REGION Network 8: WLAN5 Comm Fault
   RUNG wire#powerrail
      Contact( "reset" )
      { S7_Templates := "SrcType := USInt" } EQ_Contact(in1 := "UserDiag_HmiData".actIOSystemData.actIODeviceState[105], in2 := 3)
      wire#w1
      Coil( "DB302_HMI_Faults".SDC_Faults_0.%X5 )
   END_RUNG
   RUNG wire#powerrail
      Contact( "DB302_HMI_Faults".SDC_Faults_0.%X5 )
      I_Contact( "EMS_Fault_Reset" )
   END_RUNG wire#w1
   RUNG wire#w1
      Move(in := 6, out1 => "DB101_DB_SDC_FAULTS".SDC_Fault)
   END_RUNG
   // the same network as SCL:
   "DB302_HMI_Faults".SDC_Faults_0.%X5 := ("reset" AND ("UserDiag_HmiData".actIOSystemData.actIODeviceState[105] = 3)) OR ("DB302_HMI_Faults".SDC_Faults_0.%X5 AND NOT "EMS_Fault_Reset");
   IF "DB302_HMI_Faults".SDC_Faults_0.%X5 THEN "DB101_DB_SDC_FAULTS".SDC_Fault := 6; END_IF;
END_REGION

REGION Network 9: WLAN6 Comm Fault
   RUNG wire#powerrail
      Contact( "reset" )
      { S7_Templates := "SrcType := USInt" } EQ_Contact(in1 := "UserDiag_HmiData".actIOSystemData.actIODeviceState[106], in2 := 3)
      wire#w1
      Coil( "DB302_HMI_Faults".SDC_Faults_0.%X6 )
   END_RUNG
   RUNG wire#powerrail
      Contact( "DB302_HMI_Faults".SDC_Faults_0.%X6 )
      I_Contact( "EMS_Fault_Reset" )
   END_RUNG wire#w1
   RUNG wire#w1
      Move(in := 7, out1 => "DB101_DB_SDC_FAULTS".SDC_Fault)
   END_RUNG
   // the same network as SCL:
   "DB302_HMI_Faults".SDC_Faults_0.%X6 := ("reset" AND ("UserDiag_HmiData".actIOSystemData.actIODeviceState[106] = 3)) OR ("DB302_HMI_Faults".SDC_Faults_0.%X6 AND NOT "EMS_Fault_Reset");
   IF "DB302_HMI_Faults".SDC_Faults_0.%X6 THEN "DB101_DB_SDC_FAULTS".SDC_Fault := 7; END_IF;
END_REGION

REGION Network 10: WLAN7 Comm Fault
   RUNG wire#powerrail
      Contact( "reset" )
      { S7_Templates := "SrcType := USInt" } EQ_Contact(in1 := "UserDiag_HmiData".actIOSystemData.actIODeviceState[107], in2 := 3)
      wire#w1
      Coil( "DB302_HMI_Faults".SDC_Faults_0.%X7 )
   END_RUNG
   RUNG wire#powerrail
      Contact( "DB302_HMI_Faults".SDC_Faults_0.%X7 )
      I_Contact( "EMS_Fault_Reset" )
   END_RUNG wire#w1
   RUNG wire#w1
      Move(in := 8, out1 => "DB101_DB_SDC_FAULTS".SDC_Fault)
   END_RUNG
   // the same network as SCL:
   "DB302_HMI_Faults".SDC_Faults_0.%X7 := ("reset" AND ("UserDiag_HmiData".actIOSystemData.actIODeviceState[107] = 3)) OR ("DB302_HMI_Faults".SDC_Faults_0.%X7 AND NOT "EMS_Fault_Reset");
   IF "DB302_HMI_Faults".SDC_Faults_0.%X7 THEN "DB101_DB_SDC_FAULTS".SDC_Fault := 8; END_IF;
END_REGION

REGION Network 11: WLAN8 Comm Fault
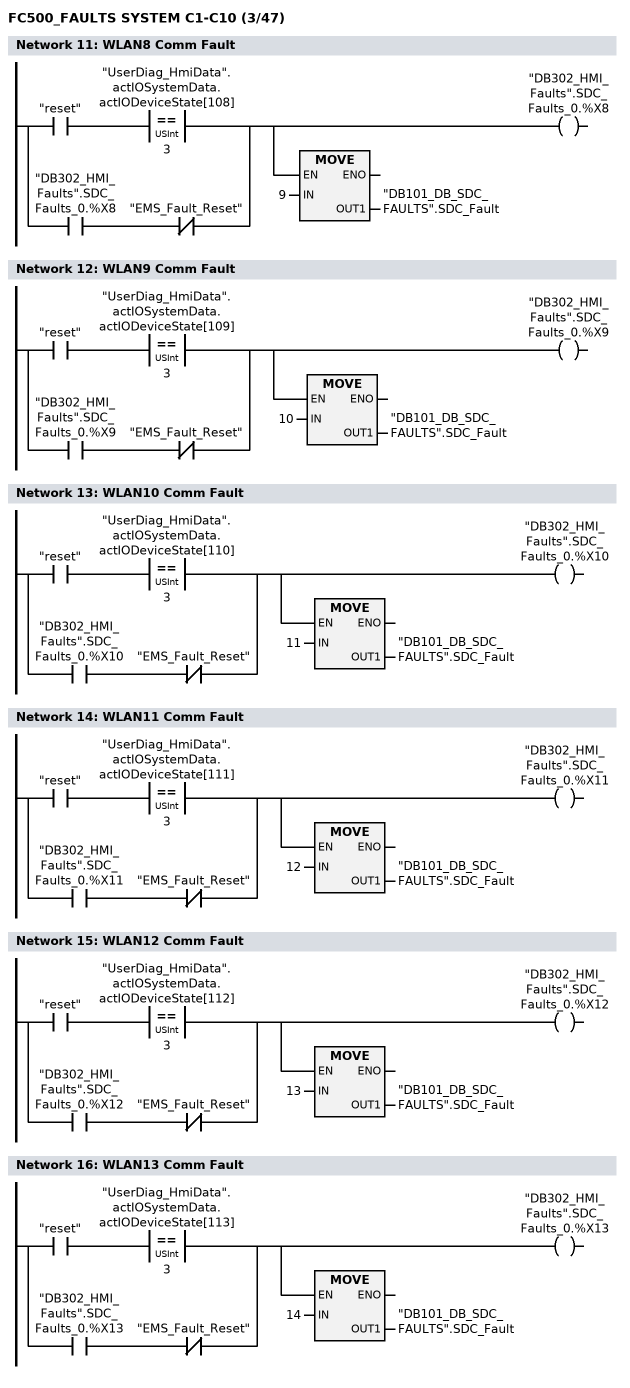
   RUNG wire#powerrail
      Contact( "reset" )
      { S7_Templates := "SrcType := USInt" } EQ_Contact(in1 := "UserDiag_HmiData".actIOSystemData.actIODeviceState[108], in2 := 3)
      wire#w1
      Coil( "DB302_HMI_Faults".SDC_Faults_0.%X8 )
   END_RUNG
   RUNG wire#powerrail
      Contact( "DB302_HMI_Faults".SDC_Faults_0.%X8 )
      I_Contact( "EMS_Fault_Reset" )
   END_RUNG wire#w1
   RUNG wire#w1
      Move(in := 9, out1 => "DB101_DB_SDC_FAULTS".SDC_Fault)
   END_RUNG
   // the same network as SCL:
   "DB302_HMI_Faults".SDC_Faults_0.%X8 := ("reset" AND ("UserDiag_HmiData".actIOSystemData.actIODeviceState[108] = 3)) OR ("DB302_HMI_Faults".SDC_Faults_0.%X8 AND NOT "EMS_Fault_Reset");
   IF "DB302_HMI_Faults".SDC_Faults_0.%X8 THEN "DB101_DB_SDC_FAULTS".SDC_Fault := 9; END_IF;
END_REGION

REGION Network 12: WLAN9 Comm Fault
   RUNG wire#powerrail
      Contact( "reset" )
      { S7_Templates := "SrcType := USInt" } EQ_Contact(in1 := "UserDiag_HmiData".actIOSystemData.actIODeviceState[109], in2 := 3)
      wire#w1
      Coil( "DB302_HMI_Faults".SDC_Faults_0.%X9 )
   END_RUNG
   RUNG wire#powerrail
      Contact( "DB302_HMI_Faults".SDC_Faults_0.%X9 )
      I_Contact( "EMS_Fault_Reset" )
   END_RUNG wire#w1
   RUNG wire#w1
      Move(in := 10, out1 => "DB101_DB_SDC_FAULTS".SDC_Fault)
   END_RUNG
   // the same network as SCL:
   "DB302_HMI_Faults".SDC_Faults_0.%X9 := ("reset" AND ("UserDiag_HmiData".actIOSystemData.actIODeviceState[109] = 3)) OR ("DB302_HMI_Faults".SDC_Faults_0.%X9 AND NOT "EMS_Fault_Reset");
   IF "DB302_HMI_Faults".SDC_Faults_0.%X9 THEN "DB101_DB_SDC_FAULTS".SDC_Fault := 10; END_IF;
END_REGION

REGION Network 13: WLAN10 Comm Fault
   RUNG wire#powerrail
      Contact( "reset" )
      { S7_Templates := "SrcType := USInt" } EQ_Contact(in1 := "UserDiag_HmiData".actIOSystemData.actIODeviceState[110], in2 := 3)
      wire#w1
      Coil( "DB302_HMI_Faults".SDC_Faults_0.%X10 )
   END_RUNG
   RUNG wire#powerrail
      Contact( "DB302_HMI_Faults".SDC_Faults_0.%X10 )
      I_Contact( "EMS_Fault_Reset" )
   END_RUNG wire#w1
   RUNG wire#w1
      Move(in := 11, out1 => "DB101_DB_SDC_FAULTS".SDC_Fault)
   END_RUNG
   // the same network as SCL:
   "DB302_HMI_Faults".SDC_Faults_0.%X10 := ("reset" AND ("UserDiag_HmiData".actIOSystemData.actIODeviceState[110] = 3)) OR ("DB302_HMI_Faults".SDC_Faults_0.%X10 AND NOT "EMS_Fault_Reset");
   IF "DB302_HMI_Faults".SDC_Faults_0.%X10 THEN "DB101_DB_SDC_FAULTS".SDC_Fault := 11; END_IF;
END_REGION

REGION Network 14: WLAN11 Comm Fault
   RUNG wire#powerrail
      Contact( "reset" )
      { S7_Templates := "SrcType := USInt" } EQ_Contact(in1 := "UserDiag_HmiData".actIOSystemData.actIODeviceState[111], in2 := 3)
      wire#w1
      Coil( "DB302_HMI_Faults".SDC_Faults_0.%X11 )
   END_RUNG
   RUNG wire#powerrail
      Contact( "DB302_HMI_Faults".SDC_Faults_0.%X11 )
      I_Contact( "EMS_Fault_Reset" )
   END_RUNG wire#w1
   RUNG wire#w1
      Move(in := 12, out1 => "DB101_DB_SDC_FAULTS".SDC_Fault)
   END_RUNG
   // the same network as SCL:
   "DB302_HMI_Faults".SDC_Faults_0.%X11 := ("reset" AND ("UserDiag_HmiData".actIOSystemData.actIODeviceState[111] = 3)) OR ("DB302_HMI_Faults".SDC_Faults_0.%X11 AND NOT "EMS_Fault_Reset");
   IF "DB302_HMI_Faults".SDC_Faults_0.%X11 THEN "DB101_DB_SDC_FAULTS".SDC_Fault := 12; END_IF;
END_REGION

REGION Network 15: WLAN12 Comm Fault
   RUNG wire#powerrail
      Contact( "reset" )
      { S7_Templates := "SrcType := USInt" } EQ_Contact(in1 := "UserDiag_HmiData".actIOSystemData.actIODeviceState[112], in2 := 3)
      wire#w1
      Coil( "DB302_HMI_Faults".SDC_Faults_0.%X12 )
   END_RUNG
   RUNG wire#powerrail
      Contact( "DB302_HMI_Faults".SDC_Faults_0.%X12 )
      I_Contact( "EMS_Fault_Reset" )
   END_RUNG wire#w1
   RUNG wire#w1
      Move(in := 13, out1 => "DB101_DB_SDC_FAULTS".SDC_Fault)
   END_RUNG
   // the same network as SCL:
   "DB302_HMI_Faults".SDC_Faults_0.%X12 := ("reset" AND ("UserDiag_HmiData".actIOSystemData.actIODeviceState[112] = 3)) OR ("DB302_HMI_Faults".SDC_Faults_0.%X12 AND NOT "EMS_Fault_Reset");
   IF "DB302_HMI_Faults".SDC_Faults_0.%X12 THEN "DB101_DB_SDC_FAULTS".SDC_Fault := 13; END_IF;
END_REGION

REGION Network 16: WLAN13 Comm Fault
   RUNG wire#powerrail
      Contact( "reset" )
      { S7_Templates := "SrcType := USInt" } EQ_Contact(in1 := "UserDiag_HmiData".actIOSystemData.actIODeviceState[113], in2 := 3)
      wire#w1
      Coil( "DB302_HMI_Faults".SDC_Faults_0.%X13 )
   END_RUNG
   RUNG wire#powerrail
      Contact( "DB302_HMI_Faults".SDC_Faults_0.%X13 )
      I_Contact( "EMS_Fault_Reset" )
   END_RUNG wire#w1
   RUNG wire#w1
      Move(in := 14, out1 => "DB101_DB_SDC_FAULTS".SDC_Fault)
   END_RUNG
   // the same network as SCL:
   "DB302_HMI_Faults".SDC_Faults_0.%X13 := ("reset" AND ("UserDiag_HmiData".actIOSystemData.actIODeviceState[113] = 3)) OR ("DB302_HMI_Faults".SDC_Faults_0.%X13 AND NOT "EMS_Fault_Reset");
   IF "DB302_HMI_Faults".SDC_Faults_0.%X13 THEN "DB101_DB_SDC_FAULTS".SDC_Fault := 14; END_IF;
END_REGION

REGION Network 17: WLAN14 Comm Fault
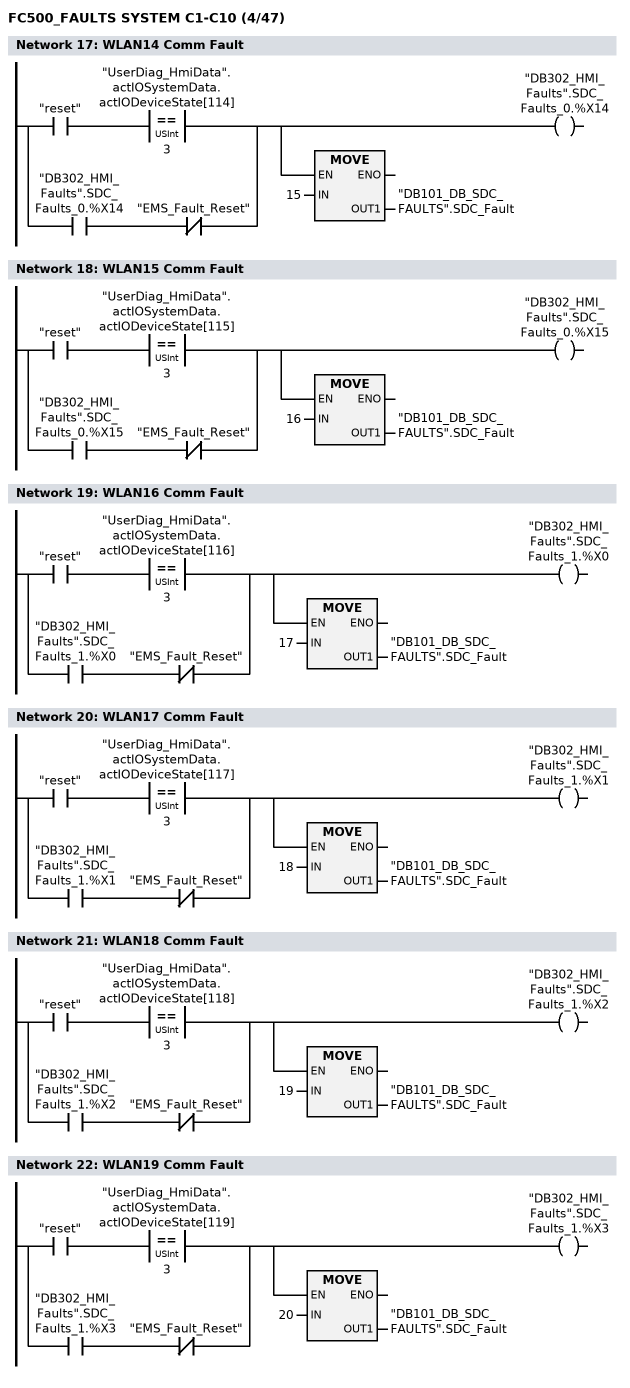
   RUNG wire#powerrail
      Contact( "reset" )
      { S7_Templates := "SrcType := USInt" } EQ_Contact(in1 := "UserDiag_HmiData".actIOSystemData.actIODeviceState[114], in2 := 3)
      wire#w1
      Coil( "DB302_HMI_Faults".SDC_Faults_0.%X14 )
   END_RUNG
   RUNG wire#powerrail
      Contact( "DB302_HMI_Faults".SDC_Faults_0.%X14 )
      I_Contact( "EMS_Fault_Reset" )
   END_RUNG wire#w1
   RUNG wire#w1
      Move(in := 15, out1 => "DB101_DB_SDC_FAULTS".SDC_Fault)
   END_RUNG
   // the same network as SCL:
   "DB302_HMI_Faults".SDC_Faults_0.%X14 := ("reset" AND ("UserDiag_HmiData".actIOSystemData.actIODeviceState[114] = 3)) OR ("DB302_HMI_Faults".SDC_Faults_0.%X14 AND NOT "EMS_Fault_Reset");
   IF "DB302_HMI_Faults".SDC_Faults_0.%X14 THEN "DB101_DB_SDC_FAULTS".SDC_Fault := 15; END_IF;
END_REGION

REGION Network 18: WLAN15 Comm Fault
   RUNG wire#powerrail
      Contact( "reset" )
      { S7_Templates := "SrcType := USInt" } EQ_Contact(in1 := "UserDiag_HmiData".actIOSystemData.actIODeviceState[115], in2 := 3)
      wire#w1
      Coil( "DB302_HMI_Faults".SDC_Faults_0.%X15 )
   END_RUNG
   RUNG wire#powerrail
      Contact( "DB302_HMI_Faults".SDC_Faults_0.%X15 )
      I_Contact( "EMS_Fault_Reset" )
   END_RUNG wire#w1
   RUNG wire#w1
      Move(in := 16, out1 => "DB101_DB_SDC_FAULTS".SDC_Fault)
   END_RUNG
   // the same network as SCL:
   "DB302_HMI_Faults".SDC_Faults_0.%X15 := ("reset" AND ("UserDiag_HmiData".actIOSystemData.actIODeviceState[115] = 3)) OR ("DB302_HMI_Faults".SDC_Faults_0.%X15 AND NOT "EMS_Fault_Reset");
   IF "DB302_HMI_Faults".SDC_Faults_0.%X15 THEN "DB101_DB_SDC_FAULTS".SDC_Fault := 16; END_IF;
END_REGION

REGION Network 19: WLAN16 Comm Fault
   RUNG wire#powerrail
      Contact( "reset" )
      { S7_Templates := "SrcType := USInt" } EQ_Contact(in1 := "UserDiag_HmiData".actIOSystemData.actIODeviceState[116], in2 := 3)
      wire#w1
      Coil( "DB302_HMI_Faults".SDC_Faults_1.%X0 )
   END_RUNG
   RUNG wire#powerrail
      Contact( "DB302_HMI_Faults".SDC_Faults_1.%X0 )
      I_Contact( "EMS_Fault_Reset" )
   END_RUNG wire#w1
   RUNG wire#w1
      Move(in := 17, out1 => "DB101_DB_SDC_FAULTS".SDC_Fault)
   END_RUNG
   // the same network as SCL:
   "DB302_HMI_Faults".SDC_Faults_1.%X0 := ("reset" AND ("UserDiag_HmiData".actIOSystemData.actIODeviceState[116] = 3)) OR ("DB302_HMI_Faults".SDC_Faults_1.%X0 AND NOT "EMS_Fault_Reset");
   IF "DB302_HMI_Faults".SDC_Faults_1.%X0 THEN "DB101_DB_SDC_FAULTS".SDC_Fault := 17; END_IF;
END_REGION

REGION Network 20: WLAN17 Comm Fault
   RUNG wire#powerrail
      Contact( "reset" )
      { S7_Templates := "SrcType := USInt" } EQ_Contact(in1 := "UserDiag_HmiData".actIOSystemData.actIODeviceState[117], in2 := 3)
      wire#w1
      Coil( "DB302_HMI_Faults".SDC_Faults_1.%X1 )
   END_RUNG
   RUNG wire#powerrail
      Contact( "DB302_HMI_Faults".SDC_Faults_1.%X1 )
      I_Contact( "EMS_Fault_Reset" )
   END_RUNG wire#w1
   RUNG wire#w1
      Move(in := 18, out1 => "DB101_DB_SDC_FAULTS".SDC_Fault)
   END_RUNG
   // the same network as SCL:
   "DB302_HMI_Faults".SDC_Faults_1.%X1 := ("reset" AND ("UserDiag_HmiData".actIOSystemData.actIODeviceState[117] = 3)) OR ("DB302_HMI_Faults".SDC_Faults_1.%X1 AND NOT "EMS_Fault_Reset");
   IF "DB302_HMI_Faults".SDC_Faults_1.%X1 THEN "DB101_DB_SDC_FAULTS".SDC_Fault := 18; END_IF;
END_REGION

REGION Network 21: WLAN18 Comm Fault
   RUNG wire#powerrail
      Contact( "reset" )
      { S7_Templates := "SrcType := USInt" } EQ_Contact(in1 := "UserDiag_HmiData".actIOSystemData.actIODeviceState[118], in2 := 3)
      wire#w1
      Coil( "DB302_HMI_Faults".SDC_Faults_1.%X2 )
   END_RUNG
   RUNG wire#powerrail
      Contact( "DB302_HMI_Faults".SDC_Faults_1.%X2 )
      I_Contact( "EMS_Fault_Reset" )
   END_RUNG wire#w1
   RUNG wire#w1
      Move(in := 19, out1 => "DB101_DB_SDC_FAULTS".SDC_Fault)
   END_RUNG
   // the same network as SCL:
   "DB302_HMI_Faults".SDC_Faults_1.%X2 := ("reset" AND ("UserDiag_HmiData".actIOSystemData.actIODeviceState[118] = 3)) OR ("DB302_HMI_Faults".SDC_Faults_1.%X2 AND NOT "EMS_Fault_Reset");
   IF "DB302_HMI_Faults".SDC_Faults_1.%X2 THEN "DB101_DB_SDC_FAULTS".SDC_Fault := 19; END_IF;
END_REGION

REGION Network 22: WLAN19 Comm Fault
   RUNG wire#powerrail
      Contact( "reset" )
      { S7_Templates := "SrcType := USInt" } EQ_Contact(in1 := "UserDiag_HmiData".actIOSystemData.actIODeviceState[119], in2 := 3)
      wire#w1
      Coil( "DB302_HMI_Faults".SDC_Faults_1.%X3 )
   END_RUNG
   RUNG wire#powerrail
      Contact( "DB302_HMI_Faults".SDC_Faults_1.%X3 )
      I_Contact( "EMS_Fault_Reset" )
   END_RUNG wire#w1
   RUNG wire#w1
      Move(in := 20, out1 => "DB101_DB_SDC_FAULTS".SDC_Fault)
   END_RUNG
   // the same network as SCL:
   "DB302_HMI_Faults".SDC_Faults_1.%X3 := ("reset" AND ("UserDiag_HmiData".actIOSystemData.actIODeviceState[119] = 3)) OR ("DB302_HMI_Faults".SDC_Faults_1.%X3 AND NOT "EMS_Fault_Reset");
   IF "DB302_HMI_Faults".SDC_Faults_1.%X3 THEN "DB101_DB_SDC_FAULTS".SDC_Fault := 20; END_IF;
END_REGION

REGION Network 23: Duplicate Carrier Fault
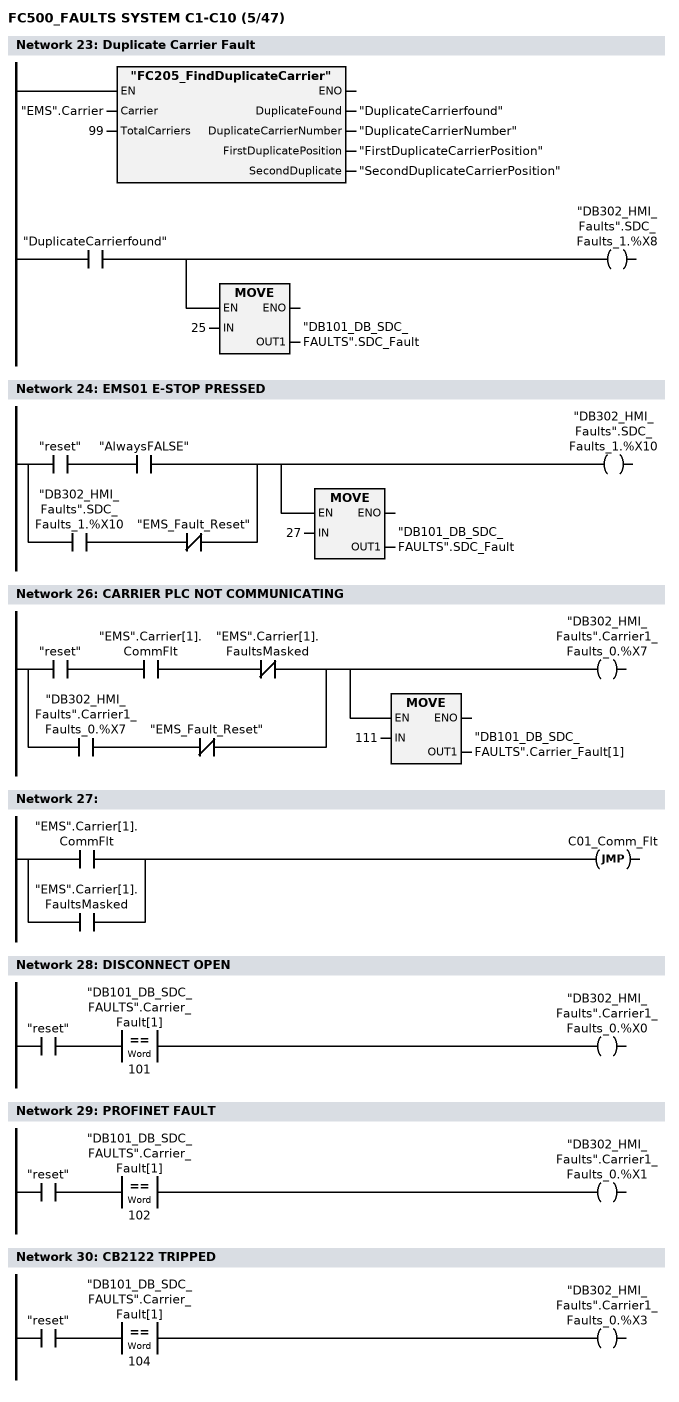
   RUNG wire#powerrail
      "FC205_FindDuplicateCarrier"(Carrier := "EMS".Carrier, TotalCarriers := 99, DuplicateFound => "DuplicateCarrierfound", DuplicateCarrierNumber => "DuplicateCarrierNumber", FirstDuplicatePosition => "FirstDuplicateCarrierPosition", SecondDuplicate => "SecondDuplicateCarrierPosition")
   END_RUNG
   RUNG wire#powerrail
      Contact( "DuplicateCarrierfound" )
      wire#w1
      Coil( "DB302_HMI_Faults".SDC_Faults_1.%X8 )
   END_RUNG
   RUNG wire#w1
      Move(in := 25, out1 => "DB101_DB_SDC_FAULTS".SDC_Fault)
   END_RUNG
   // the same network as SCL:
   "FC205_FindDuplicateCarrier"(Carrier := "EMS".Carrier,
                           TotalCarriers := 99,
                           DuplicateFound => "DuplicateCarrierfound",
                           DuplicateCarrierNumber => "DuplicateCarrierNumber",
                           FirstDuplicatePosition => "FirstDuplicateCarrierPosition",
                           SecondDuplicate => "SecondDuplicateCarrierPosition");
   "DB302_HMI_Faults".SDC_Faults_1.%X8 := "DuplicateCarrierfound";
   IF "DuplicateCarrierfound" THEN "DB101_DB_SDC_FAULTS".SDC_Fault := 25; END_IF;
END_REGION

REGION Network 24: EMS01 E-STOP PRESSED
   RUNG wire#powerrail
      Contact( "reset" )
      Contact( "AlwaysFALSE" )
      wire#w1
      Coil( "DB302_HMI_Faults".SDC_Faults_1.%X10 )
   END_RUNG
   RUNG wire#powerrail
      Contact( "DB302_HMI_Faults".SDC_Faults_1.%X10 )
      I_Contact( "EMS_Fault_Reset" )
   END_RUNG wire#w1
   RUNG wire#w1
      Move(in := 27, out1 => "DB101_DB_SDC_FAULTS".SDC_Fault)
   END_RUNG
   // the same network as SCL:
   "DB302_HMI_Faults".SDC_Faults_1.%X10 := ("reset" AND "AlwaysFALSE") OR ("DB302_HMI_Faults".SDC_Faults_1.%X10 AND NOT "EMS_Fault_Reset");
   IF "DB302_HMI_Faults".SDC_Faults_1.%X10 THEN "DB101_DB_SDC_FAULTS".SDC_Fault := 27; END_IF;
END_REGION

REGION Network 25: CARRIER 1 FAULTS
END_REGION

REGION Network 26: CARRIER PLC NOT COMMUNICATING
   RUNG wire#powerrail
      Contact( "reset" )
      Contact( "EMS".Carrier[1].CommFlt )
      I_Contact( "EMS".Carrier[1].FaultsMasked )
      wire#w1
      Coil( "DB302_HMI_Faults".Carrier1_Faults_0.%X7 )
   END_RUNG
   RUNG wire#powerrail
      Contact( "DB302_HMI_Faults".Carrier1_Faults_0.%X7 )
      I_Contact( "EMS_Fault_Reset" )
   END_RUNG wire#w1
   RUNG wire#w1
      Move(in := 111, out1 => "DB101_DB_SDC_FAULTS".Carrier_Fault[1])
   END_RUNG
   // the same network as SCL:
   "DB302_HMI_Faults".Carrier1_Faults_0.%X7 := ("reset" AND "EMS".Carrier[1].CommFlt AND NOT "EMS".Carrier[1].FaultsMasked) OR ("DB302_HMI_Faults".Carrier1_Faults_0.%X7 AND NOT "EMS_Fault_Reset");
   IF "DB302_HMI_Faults".Carrier1_Faults_0.%X7 THEN "DB101_DB_SDC_FAULTS".Carrier_Fault[1] := 111; END_IF;
END_REGION

REGION Network 27
   RUNG wire#powerrail
      Contact( "EMS".Carrier[1].CommFlt )
      wire#w1
      JumpCoil( C01_Comm_Flt )
   END_RUNG
   RUNG wire#powerrail
      Contact( "EMS".Carrier[1].FaultsMasked )
   END_RUNG wire#w1
   // the same network as SCL:
   IF "EMS".Carrier[1].CommFlt OR "EMS".Carrier[1].FaultsMasked THEN GOTO C01_Comm_Flt; END_IF;
END_REGION

REGION Network 28: DISCONNECT OPEN
   RUNG wire#powerrail
      Contact( "reset" )
      { S7_Templates := "SrcType := Word" } EQ_Contact(in1 := "DB101_DB_SDC_FAULTS".Carrier_Fault[1], in2 := 101)
      Coil( "DB302_HMI_Faults".Carrier1_Faults_0.%X0 )
   END_RUNG
   // the same network as SCL:
   "DB302_HMI_Faults".Carrier1_Faults_0.%X0 := "reset" AND ("DB101_DB_SDC_FAULTS".Carrier_Fault[1] = 101);
END_REGION

REGION Network 29: PROFINET FAULT
   RUNG wire#powerrail
      Contact( "reset" )
      { S7_Templates := "SrcType := Word" } EQ_Contact(in1 := "DB101_DB_SDC_FAULTS".Carrier_Fault[1], in2 := 102)
      Coil( "DB302_HMI_Faults".Carrier1_Faults_0.%X1 )
   END_RUNG
   // the same network as SCL:
   "DB302_HMI_Faults".Carrier1_Faults_0.%X1 := "reset" AND ("DB101_DB_SDC_FAULTS".Carrier_Fault[1] = 102);
END_REGION

REGION Network 30: CB2122 TRIPPED
   RUNG wire#powerrail
      Contact( "reset" )
      { S7_Templates := "SrcType := Word" } EQ_Contact(in1 := "DB101_DB_SDC_FAULTS".Carrier_Fault[1], in2 := 104)
      Coil( "DB302_HMI_Faults".Carrier1_Faults_0.%X3 )
   END_RUNG
   // the same network as SCL:
   "DB302_HMI_Faults".Carrier1_Faults_0.%X3 := "reset" AND ("DB101_DB_SDC_FAULTS".Carrier_Fault[1] = 104);
END_REGION

REGION Network 31: CB2123 TRIPPED
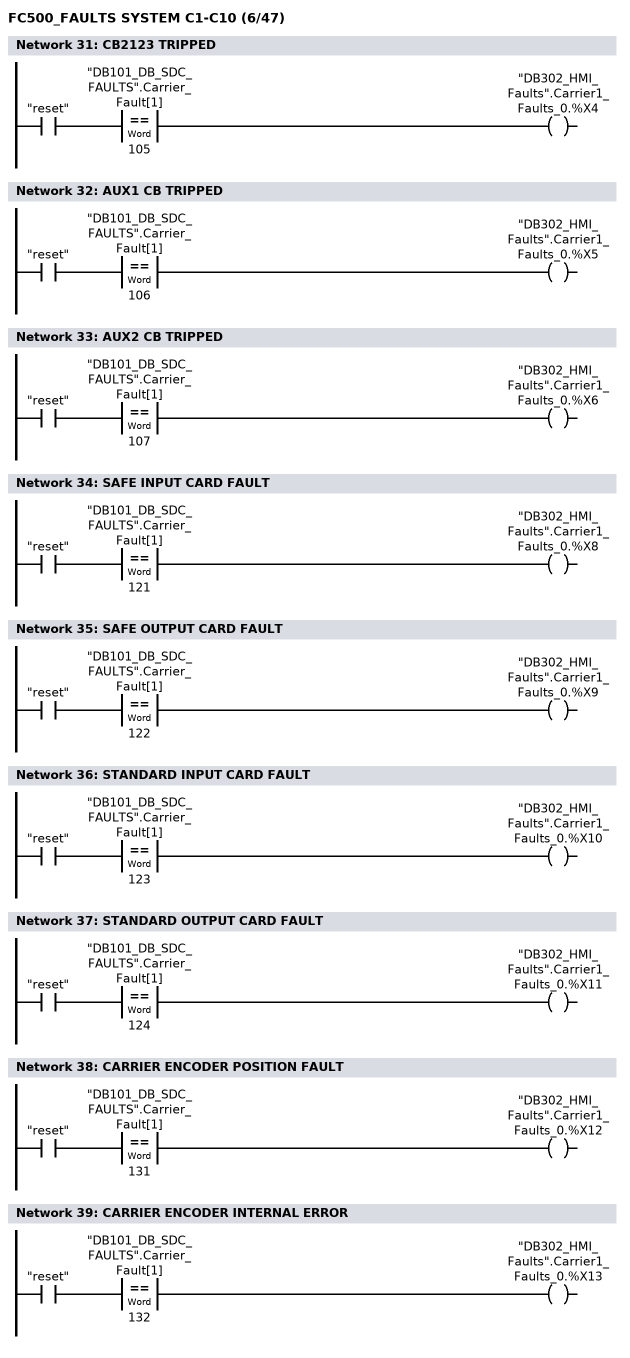
   RUNG wire#powerrail
      Contact( "reset" )
      { S7_Templates := "SrcType := Word" } EQ_Contact(in1 := "DB101_DB_SDC_FAULTS".Carrier_Fault[1], in2 := 105)
      Coil( "DB302_HMI_Faults".Carrier1_Faults_0.%X4 )
   END_RUNG
   // the same network as SCL:
   "DB302_HMI_Faults".Carrier1_Faults_0.%X4 := "reset" AND ("DB101_DB_SDC_FAULTS".Carrier_Fault[1] = 105);
END_REGION

REGION Network 32: AUX1 CB TRIPPED
   RUNG wire#powerrail
      Contact( "reset" )
      { S7_Templates := "SrcType := Word" } EQ_Contact(in1 := "DB101_DB_SDC_FAULTS".Carrier_Fault[1], in2 := 106)
      Coil( "DB302_HMI_Faults".Carrier1_Faults_0.%X5 )
   END_RUNG
   // the same network as SCL:
   "DB302_HMI_Faults".Carrier1_Faults_0.%X5 := "reset" AND ("DB101_DB_SDC_FAULTS".Carrier_Fault[1] = 106);
END_REGION

REGION Network 33: AUX2 CB TRIPPED
   RUNG wire#powerrail
      Contact( "reset" )
      { S7_Templates := "SrcType := Word" } EQ_Contact(in1 := "DB101_DB_SDC_FAULTS".Carrier_Fault[1], in2 := 107)
      Coil( "DB302_HMI_Faults".Carrier1_Faults_0.%X6 )
   END_RUNG
   // the same network as SCL:
   "DB302_HMI_Faults".Carrier1_Faults_0.%X6 := "reset" AND ("DB101_DB_SDC_FAULTS".Carrier_Fault[1] = 107);
END_REGION

REGION Network 34: SAFE INPUT CARD FAULT
   RUNG wire#powerrail
      Contact( "reset" )
      { S7_Templates := "SrcType := Word" } EQ_Contact(in1 := "DB101_DB_SDC_FAULTS".Carrier_Fault[1], in2 := 121)
      Coil( "DB302_HMI_Faults".Carrier1_Faults_0.%X8 )
   END_RUNG
   // the same network as SCL:
   "DB302_HMI_Faults".Carrier1_Faults_0.%X8 := "reset" AND ("DB101_DB_SDC_FAULTS".Carrier_Fault[1] = 121);
END_REGION

REGION Network 35: SAFE OUTPUT CARD FAULT
   RUNG wire#powerrail
      Contact( "reset" )
      { S7_Templates := "SrcType := Word" } EQ_Contact(in1 := "DB101_DB_SDC_FAULTS".Carrier_Fault[1], in2 := 122)
      Coil( "DB302_HMI_Faults".Carrier1_Faults_0.%X9 )
   END_RUNG
   // the same network as SCL:
   "DB302_HMI_Faults".Carrier1_Faults_0.%X9 := "reset" AND ("DB101_DB_SDC_FAULTS".Carrier_Fault[1] = 122);
END_REGION

REGION Network 36: STANDARD INPUT CARD FAULT
   RUNG wire#powerrail
      Contact( "reset" )
      { S7_Templates := "SrcType := Word" } EQ_Contact(in1 := "DB101_DB_SDC_FAULTS".Carrier_Fault[1], in2 := 123)
      Coil( "DB302_HMI_Faults".Carrier1_Faults_0.%X10 )
   END_RUNG
   // the same network as SCL:
   "DB302_HMI_Faults".Carrier1_Faults_0.%X10 := "reset" AND ("DB101_DB_SDC_FAULTS".Carrier_Fault[1] = 123);
END_REGION

REGION Network 37: STANDARD OUTPUT CARD FAULT
   RUNG wire#powerrail
      Contact( "reset" )
      { S7_Templates := "SrcType := Word" } EQ_Contact(in1 := "DB101_DB_SDC_FAULTS".Carrier_Fault[1], in2 := 124)
      Coil( "DB302_HMI_Faults".Carrier1_Faults_0.%X11 )
   END_RUNG
   // the same network as SCL:
   "DB302_HMI_Faults".Carrier1_Faults_0.%X11 := "reset" AND ("DB101_DB_SDC_FAULTS".Carrier_Fault[1] = 124);
END_REGION

REGION Network 38: CARRIER ENCODER POSITION FAULT
   RUNG wire#powerrail
      Contact( "reset" )
      { S7_Templates := "SrcType := Word" } EQ_Contact(in1 := "DB101_DB_SDC_FAULTS".Carrier_Fault[1], in2 := 131)
      Coil( "DB302_HMI_Faults".Carrier1_Faults_0.%X12 )
   END_RUNG
   // the same network as SCL:
   "DB302_HMI_Faults".Carrier1_Faults_0.%X12 := "reset" AND ("DB101_DB_SDC_FAULTS".Carrier_Fault[1] = 131);
END_REGION

REGION Network 39: CARRIER ENCODER INTERNAL ERROR
   RUNG wire#powerrail
      Contact( "reset" )
      { S7_Templates := "SrcType := Word" } EQ_Contact(in1 := "DB101_DB_SDC_FAULTS".Carrier_Fault[1], in2 := 132)
      Coil( "DB302_HMI_Faults".Carrier1_Faults_0.%X13 )
   END_RUNG
   // the same network as SCL:
   "DB302_HMI_Faults".Carrier1_Faults_0.%X13 := "reset" AND ("DB101_DB_SDC_FAULTS".Carrier_Fault[1] = 132);
END_REGION

REGION Network 40: CARRIER ENCODER COMM FAULT
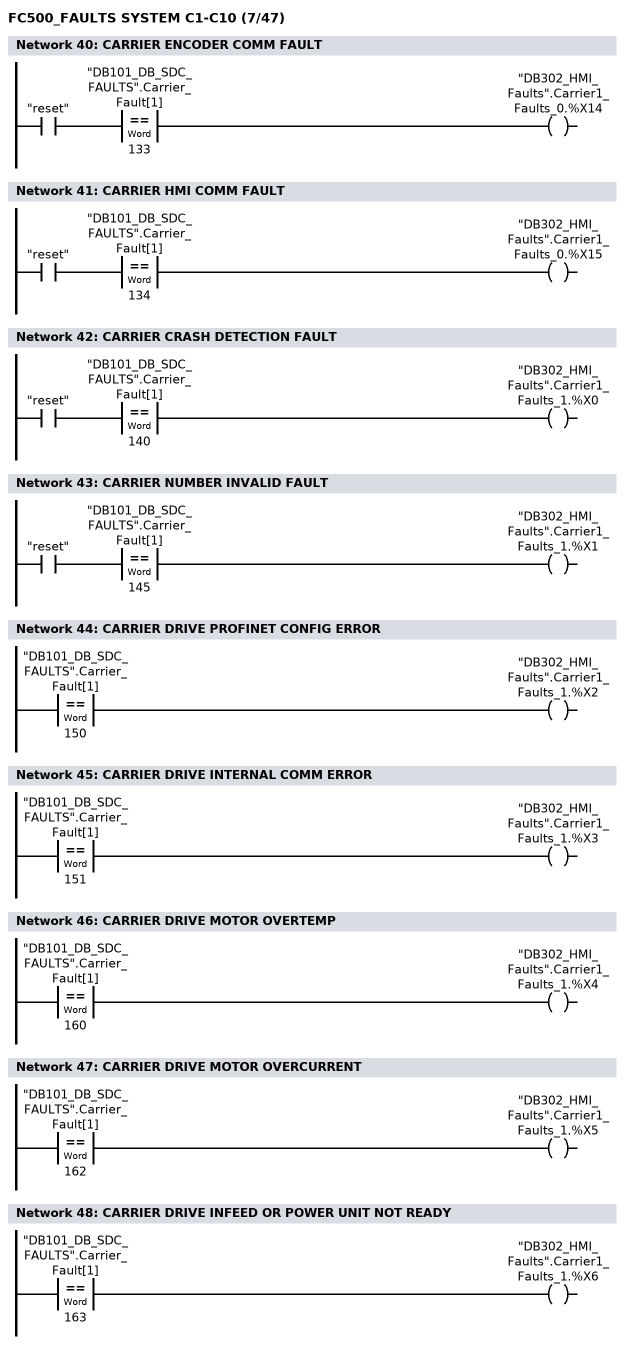
   RUNG wire#powerrail
      Contact( "reset" )
      { S7_Templates := "SrcType := Word" } EQ_Contact(in1 := "DB101_DB_SDC_FAULTS".Carrier_Fault[1], in2 := 133)
      Coil( "DB302_HMI_Faults".Carrier1_Faults_0.%X14 )
   END_RUNG
   // the same network as SCL:
   "DB302_HMI_Faults".Carrier1_Faults_0.%X14 := "reset" AND ("DB101_DB_SDC_FAULTS".Carrier_Fault[1] = 133);
END_REGION

REGION Network 41: CARRIER HMI COMM FAULT
   RUNG wire#powerrail
      Contact( "reset" )
      { S7_Templates := "SrcType := Word" } EQ_Contact(in1 := "DB101_DB_SDC_FAULTS".Carrier_Fault[1], in2 := 134)
      Coil( "DB302_HMI_Faults".Carrier1_Faults_0.%X15 )
   END_RUNG
   // the same network as SCL:
   "DB302_HMI_Faults".Carrier1_Faults_0.%X15 := "reset" AND ("DB101_DB_SDC_FAULTS".Carrier_Fault[1] = 134);
END_REGION

REGION Network 42: CARRIER CRASH DETECTION FAULT
   RUNG wire#powerrail
      Contact( "reset" )
      { S7_Templates := "SrcType := Word" } EQ_Contact(in1 := "DB101_DB_SDC_FAULTS".Carrier_Fault[1], in2 := 140)
      Coil( "DB302_HMI_Faults".Carrier1_Faults_1.%X0 )
   END_RUNG
   // the same network as SCL:
   "DB302_HMI_Faults".Carrier1_Faults_1.%X0 := "reset" AND ("DB101_DB_SDC_FAULTS".Carrier_Fault[1] = 140);
END_REGION

REGION Network 43: CARRIER NUMBER INVALID FAULT
   RUNG wire#powerrail
      Contact( "reset" )
      { S7_Templates := "SrcType := Word" } EQ_Contact(in1 := "DB101_DB_SDC_FAULTS".Carrier_Fault[1], in2 := 145)
      Coil( "DB302_HMI_Faults".Carrier1_Faults_1.%X1 )
   END_RUNG
   // the same network as SCL:
   "DB302_HMI_Faults".Carrier1_Faults_1.%X1 := "reset" AND ("DB101_DB_SDC_FAULTS".Carrier_Fault[1] = 145);
END_REGION

REGION Network 44: CARRIER DRIVE PROFINET CONFIG ERROR
   RUNG wire#powerrail
      { S7_Templates := "SrcType := Word" } EQ_Contact(in1 := "DB101_DB_SDC_FAULTS".Carrier_Fault[1], in2 := 150)
      Coil( "DB302_HMI_Faults".Carrier1_Faults_1.%X2 )
   END_RUNG
   // the same network as SCL:
   "DB302_HMI_Faults".Carrier1_Faults_1.%X2 := "DB101_DB_SDC_FAULTS".Carrier_Fault[1] = 150;
END_REGION

REGION Network 45: CARRIER DRIVE INTERNAL COMM ERROR
   RUNG wire#powerrail
      { S7_Templates := "SrcType := Word" } EQ_Contact(in1 := "DB101_DB_SDC_FAULTS".Carrier_Fault[1], in2 := 151)
      Coil( "DB302_HMI_Faults".Carrier1_Faults_1.%X3 )
   END_RUNG
   // the same network as SCL:
   "DB302_HMI_Faults".Carrier1_Faults_1.%X3 := "DB101_DB_SDC_FAULTS".Carrier_Fault[1] = 151;
END_REGION

REGION Network 46: CARRIER DRIVE MOTOR OVERTEMP
   RUNG wire#powerrail
      { S7_Templates := "SrcType := Word" } EQ_Contact(in1 := "DB101_DB_SDC_FAULTS".Carrier_Fault[1], in2 := 160)
      Coil( "DB302_HMI_Faults".Carrier1_Faults_1.%X4 )
   END_RUNG
   // the same network as SCL:
   "DB302_HMI_Faults".Carrier1_Faults_1.%X4 := "DB101_DB_SDC_FAULTS".Carrier_Fault[1] = 160;
END_REGION

REGION Network 47: CARRIER DRIVE MOTOR OVERCURRENT
   RUNG wire#powerrail
      { S7_Templates := "SrcType := Word" } EQ_Contact(in1 := "DB101_DB_SDC_FAULTS".Carrier_Fault[1], in2 := 162)
      Coil( "DB302_HMI_Faults".Carrier1_Faults_1.%X5 )
   END_RUNG
   // the same network as SCL:
   "DB302_HMI_Faults".Carrier1_Faults_1.%X5 := "DB101_DB_SDC_FAULTS".Carrier_Fault[1] = 162;
END_REGION

REGION Network 48: CARRIER DRIVE INFEED OR POWER UNIT NOT READY
   RUNG wire#powerrail
      { S7_Templates := "SrcType := Word" } EQ_Contact(in1 := "DB101_DB_SDC_FAULTS".Carrier_Fault[1], in2 := 163)
      Coil( "DB302_HMI_Faults".Carrier1_Faults_1.%X6 )
   END_RUNG
   // the same network as SCL:
   "DB302_HMI_Faults".Carrier1_Faults_1.%X6 := "DB101_DB_SDC_FAULTS".Carrier_Fault[1] = 163;
END_REGION

REGION Network 49: CARRIER DRIVE SHORT CIRCUIT / GROUND FAULT DETECTED
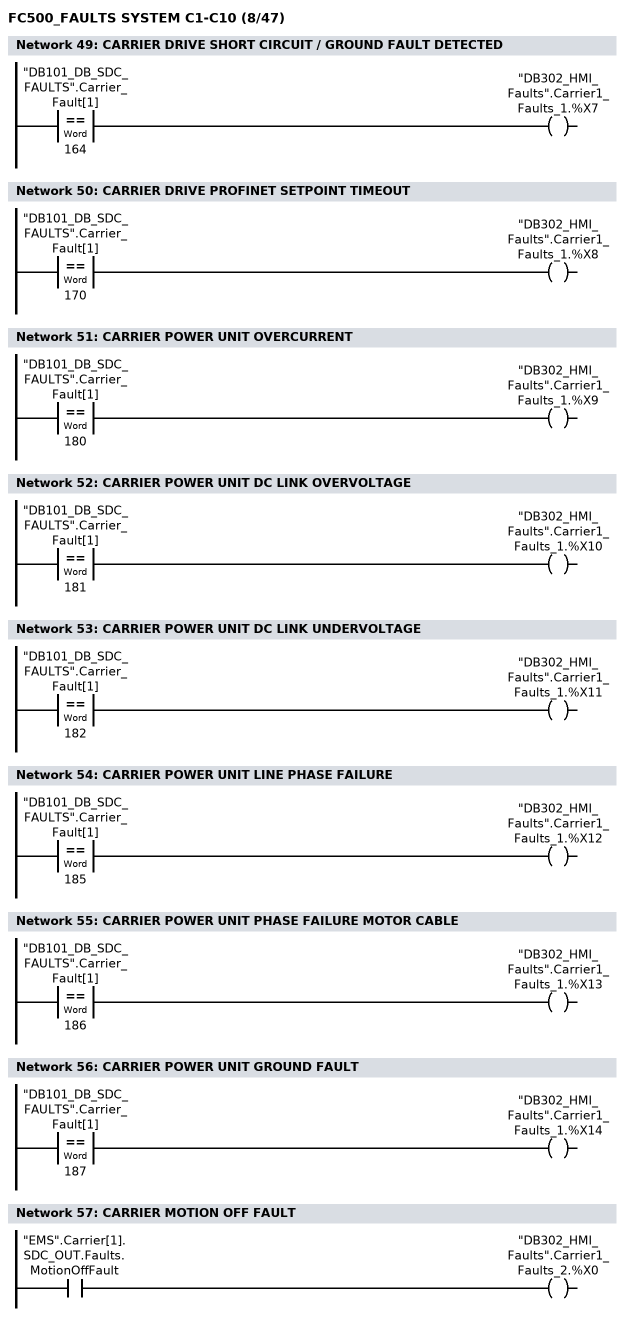
   RUNG wire#powerrail
      { S7_Templates := "SrcType := Word" } EQ_Contact(in1 := "DB101_DB_SDC_FAULTS".Carrier_Fault[1], in2 := 164)
      Coil( "DB302_HMI_Faults".Carrier1_Faults_1.%X7 )
   END_RUNG
   // the same network as SCL:
   "DB302_HMI_Faults".Carrier1_Faults_1.%X7 := "DB101_DB_SDC_FAULTS".Carrier_Fault[1] = 164;
END_REGION

REGION Network 50: CARRIER DRIVE PROFINET SETPOINT TIMEOUT
   RUNG wire#powerrail
      { S7_Templates := "SrcType := Word" } EQ_Contact(in1 := "DB101_DB_SDC_FAULTS".Carrier_Fault[1], in2 := 170)
      Coil( "DB302_HMI_Faults".Carrier1_Faults_1.%X8 )
   END_RUNG
   // the same network as SCL:
   "DB302_HMI_Faults".Carrier1_Faults_1.%X8 := "DB101_DB_SDC_FAULTS".Carrier_Fault[1] = 170;
END_REGION

REGION Network 51: CARRIER POWER UNIT OVERCURRENT
   RUNG wire#powerrail
      { S7_Templates := "SrcType := Word" } EQ_Contact(in1 := "DB101_DB_SDC_FAULTS".Carrier_Fault[1], in2 := 180)
      Coil( "DB302_HMI_Faults".Carrier1_Faults_1.%X9 )
   END_RUNG
   // the same network as SCL:
   "DB302_HMI_Faults".Carrier1_Faults_1.%X9 := "DB101_DB_SDC_FAULTS".Carrier_Fault[1] = 180;
END_REGION

REGION Network 52: CARRIER POWER UNIT DC LINK OVERVOLTAGE
   RUNG wire#powerrail
      { S7_Templates := "SrcType := Word" } EQ_Contact(in1 := "DB101_DB_SDC_FAULTS".Carrier_Fault[1], in2 := 181)
      Coil( "DB302_HMI_Faults".Carrier1_Faults_1.%X10 )
   END_RUNG
   // the same network as SCL:
   "DB302_HMI_Faults".Carrier1_Faults_1.%X10 := "DB101_DB_SDC_FAULTS".Carrier_Fault[1] = 181;
END_REGION

REGION Network 53: CARRIER POWER UNIT DC LINK UNDERVOLTAGE
   RUNG wire#powerrail
      { S7_Templates := "SrcType := Word" } EQ_Contact(in1 := "DB101_DB_SDC_FAULTS".Carrier_Fault[1], in2 := 182)
      Coil( "DB302_HMI_Faults".Carrier1_Faults_1.%X11 )
   END_RUNG
   // the same network as SCL:
   "DB302_HMI_Faults".Carrier1_Faults_1.%X11 := "DB101_DB_SDC_FAULTS".Carrier_Fault[1] = 182;
END_REGION

REGION Network 54: CARRIER POWER UNIT LINE PHASE FAILURE
   RUNG wire#powerrail
      { S7_Templates := "SrcType := Word" } EQ_Contact(in1 := "DB101_DB_SDC_FAULTS".Carrier_Fault[1], in2 := 185)
      Coil( "DB302_HMI_Faults".Carrier1_Faults_1.%X12 )
   END_RUNG
   // the same network as SCL:
   "DB302_HMI_Faults".Carrier1_Faults_1.%X12 := "DB101_DB_SDC_FAULTS".Carrier_Fault[1] = 185;
END_REGION

REGION Network 55: CARRIER POWER UNIT PHASE FAILURE MOTOR CABLE
   RUNG wire#powerrail
      { S7_Templates := "SrcType := Word" } EQ_Contact(in1 := "DB101_DB_SDC_FAULTS".Carrier_Fault[1], in2 := 186)
      Coil( "DB302_HMI_Faults".Carrier1_Faults_1.%X13 )
   END_RUNG
   // the same network as SCL:
   "DB302_HMI_Faults".Carrier1_Faults_1.%X13 := "DB101_DB_SDC_FAULTS".Carrier_Fault[1] = 186;
END_REGION

REGION Network 56: CARRIER POWER UNIT GROUND FAULT
   RUNG wire#powerrail
      { S7_Templates := "SrcType := Word" } EQ_Contact(in1 := "DB101_DB_SDC_FAULTS".Carrier_Fault[1], in2 := 187)
      Coil( "DB302_HMI_Faults".Carrier1_Faults_1.%X14 )
   END_RUNG
   // the same network as SCL:
   "DB302_HMI_Faults".Carrier1_Faults_1.%X14 := "DB101_DB_SDC_FAULTS".Carrier_Fault[1] = 187;
END_REGION

REGION Network 57: CARRIER MOTION OFF FAULT
   RUNG wire#powerrail
      Contact( "EMS".Carrier[1].SDC_OUT.Faults.MotionOffFault )
      Coil( "DB302_HMI_Faults".Carrier1_Faults_2.%X0 )
   END_RUNG
   // the same network as SCL:
   "DB302_HMI_Faults".Carrier1_Faults_2.%X0 := "EMS".Carrier[1].SDC_OUT.Faults.MotionOffFault;
END_REGION

REGION Network 58: CARRIER MOTION ON FAULT
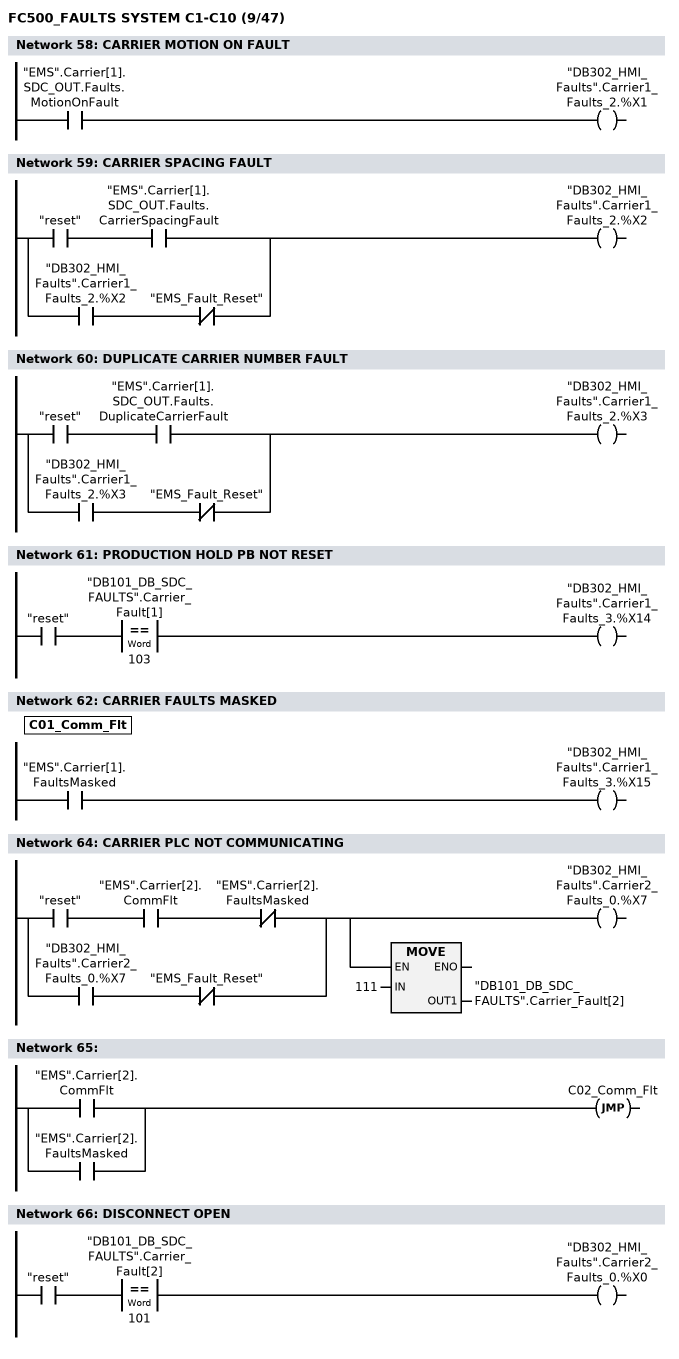
   RUNG wire#powerrail
      Contact( "EMS".Carrier[1].SDC_OUT.Faults.MotionOnFault )
      Coil( "DB302_HMI_Faults".Carrier1_Faults_2.%X1 )
   END_RUNG
   // the same network as SCL:
   "DB302_HMI_Faults".Carrier1_Faults_2.%X1 := "EMS".Carrier[1].SDC_OUT.Faults.MotionOnFault;
END_REGION

REGION Network 59: CARRIER SPACING FAULT
   RUNG wire#powerrail
      Contact( "reset" )
      Contact( "EMS".Carrier[1].SDC_OUT.Faults.CarrierSpacingFault )
      wire#w1
      Coil( "DB302_HMI_Faults".Carrier1_Faults_2.%X2 )
   END_RUNG
   RUNG wire#powerrail
      Contact( "DB302_HMI_Faults".Carrier1_Faults_2.%X2 )
      I_Contact( "EMS_Fault_Reset" )
   END_RUNG wire#w1
   // the same network as SCL:
   "DB302_HMI_Faults".Carrier1_Faults_2.%X2 := ("reset" AND "EMS".Carrier[1].SDC_OUT.Faults.CarrierSpacingFault) OR ("DB302_HMI_Faults".Carrier1_Faults_2.%X2 AND NOT "EMS_Fault_Reset");
END_REGION

REGION Network 60: DUPLICATE CARRIER NUMBER FAULT
   RUNG wire#powerrail
      Contact( "reset" )
      Contact( "EMS".Carrier[1].SDC_OUT.Faults.DuplicateCarrierFault )
      wire#w1
      Coil( "DB302_HMI_Faults".Carrier1_Faults_2.%X3 )
   END_RUNG
   RUNG wire#powerrail
      Contact( "DB302_HMI_Faults".Carrier1_Faults_2.%X3 )
      I_Contact( "EMS_Fault_Reset" )
   END_RUNG wire#w1
   // the same network as SCL:
   "DB302_HMI_Faults".Carrier1_Faults_2.%X3 := ("reset" AND "EMS".Carrier[1].SDC_OUT.Faults.DuplicateCarrierFault) OR ("DB302_HMI_Faults".Carrier1_Faults_2.%X3 AND NOT "EMS_Fault_Reset");
END_REGION

REGION Network 61: PRODUCTION HOLD PB NOT RESET
   RUNG wire#powerrail
      Contact( "reset" )
      { S7_Templates := "SrcType := Word" } EQ_Contact(in1 := "DB101_DB_SDC_FAULTS".Carrier_Fault[1], in2 := 103)
      Coil( "DB302_HMI_Faults".Carrier1_Faults_3.%X14 )
   END_RUNG
   // the same network as SCL:
   "DB302_HMI_Faults".Carrier1_Faults_3.%X14 := "reset" AND ("DB101_DB_SDC_FAULTS".Carrier_Fault[1] = 103);
END_REGION

REGION Network 62: CARRIER FAULTS MASKED
   Label( C01_Comm_Flt )
   RUNG wire#powerrail
      Contact( "EMS".Carrier[1].FaultsMasked )
      Coil( "DB302_HMI_Faults".Carrier1_Faults_3.%X15 )
   END_RUNG
   // the same network as SCL:
   C01_Comm_Flt:
   "DB302_HMI_Faults".Carrier1_Faults_3.%X15 := "EMS".Carrier[1].FaultsMasked;
END_REGION

REGION Network 63: Carrier 2 Faults
END_REGION

REGION Network 64: CARRIER PLC NOT COMMUNICATING
   RUNG wire#powerrail
      Contact( "reset" )
      Contact( "EMS".Carrier[2].CommFlt )
      I_Contact( "EMS".Carrier[2].FaultsMasked )
      wire#w1
      Coil( "DB302_HMI_Faults".Carrier2_Faults_0.%X7 )
   END_RUNG
   RUNG wire#powerrail
      Contact( "DB302_HMI_Faults".Carrier2_Faults_0.%X7 )
      I_Contact( "EMS_Fault_Reset" )
   END_RUNG wire#w1
   RUNG wire#w1
      Move(in := 111, out1 => "DB101_DB_SDC_FAULTS".Carrier_Fault[2])
   END_RUNG
   // the same network as SCL:
   "DB302_HMI_Faults".Carrier2_Faults_0.%X7 := ("reset" AND "EMS".Carrier[2].CommFlt AND NOT "EMS".Carrier[2].FaultsMasked) OR ("DB302_HMI_Faults".Carrier2_Faults_0.%X7 AND NOT "EMS_Fault_Reset");
   IF "DB302_HMI_Faults".Carrier2_Faults_0.%X7 THEN "DB101_DB_SDC_FAULTS".Carrier_Fault[2] := 111; END_IF;
END_REGION

REGION Network 65
   RUNG wire#powerrail
      Contact( "EMS".Carrier[2].CommFlt )
      wire#w1
      JumpCoil( C02_Comm_Flt )
   END_RUNG
   RUNG wire#powerrail
      Contact( "EMS".Carrier[2].FaultsMasked )
   END_RUNG wire#w1
   // the same network as SCL:
   IF "EMS".Carrier[2].CommFlt OR "EMS".Carrier[2].FaultsMasked THEN GOTO C02_Comm_Flt; END_IF;
END_REGION

REGION Network 66: DISCONNECT OPEN
   RUNG wire#powerrail
      Contact( "reset" )
      { S7_Templates := "SrcType := Word" } EQ_Contact(in1 := "DB101_DB_SDC_FAULTS".Carrier_Fault[2], in2 := 101)
      Coil( "DB302_HMI_Faults".Carrier2_Faults_0.%X0 )
   END_RUNG
   // the same network as SCL:
   "DB302_HMI_Faults".Carrier2_Faults_0.%X0 := "reset" AND ("DB101_DB_SDC_FAULTS".Carrier_Fault[2] = 101);
END_REGION

REGION Network 67: PROFINET FAULT
